REGION Network 29: a | b | c | d | e |
   RUNG wire#powerrail
      I_Contact( #DONE )
      { S7_Templates := "SrcType := WChar" } EQ_Contact(in1 := #UNICODE, in2 := WCHAR#'a')
      Move(in := 16#61, out1 => #ASCII_HEX)
      S_Coil( #DONE )
   END_RUNG
   RUNG wire#powerrail
      I_Contact( #DONE )
      { S7_Templates := "SrcType := WChar" } EQ_Contact(in1 := #UNICODE, in2 := WCHAR#'b')
      Move(in := 16#62, out1 => #ASCII_HEX)
      S_Coil( #DONE )
   END_RUNG
   RUNG wire#powerrail
      I_Contact( #DONE )
      { S7_Templates := "SrcType := WChar" } EQ_Contact(in1 := #UNICODE, in2 := WCHAR#'c')
      Move(in := 16#63, out1 => #ASCII_HEX)
      S_Coil( #DONE )
   END_RUNG
   RUNG wire#powerrail
      I_Contact( #DONE )
      { S7_Templates := "SrcType := WChar" } EQ_Contact(in1 := #UNICODE, in2 := WCHAR#'d')
      Move(in := 16#64, out1 => #ASCII_HEX)
      S_Coil( #DONE )
   END_RUNG
   RUNG wire#powerrail
      I_Contact( #DONE )
      { S7_Templates := "SrcType := WChar" } EQ_Contact(in1 := #UNICODE, in2 := WCHAR#'e')
      Move(in := 16#65, out1 => #ASCII_HEX)
      S_Coil( #DONE )
   END_RUNG
   // the same network as SCL:
   IF NOT #DONE AND (#UNICODE = WCHAR#'a') THEN
       #ASCII_HEX := 16#61;
       #DONE := TRUE;
   END_IF;
   IF NOT #DONE AND (#UNICODE = WCHAR#'b') THEN
       #ASCII_HEX := 16#62;
       #DONE := TRUE;
   END_IF;
   IF NOT #DONE AND (#UNICODE = WCHAR#'c') THEN
       #ASCII_HEX := 16#63;
       #DONE := TRUE;
   END_IF;
   IF NOT #DONE AND (#UNICODE = WCHAR#'d') THEN
       #ASCII_HEX := 16#64;
       #DONE := TRUE;
   END_IF;
   IF NOT #DONE AND (#UNICODE = WCHAR#'e') THEN
       #ASCII_HEX := 16#65;
       #DONE := TRUE;
   END_IF;
END_REGION

REGION Network 30: f | g | h | i | j |
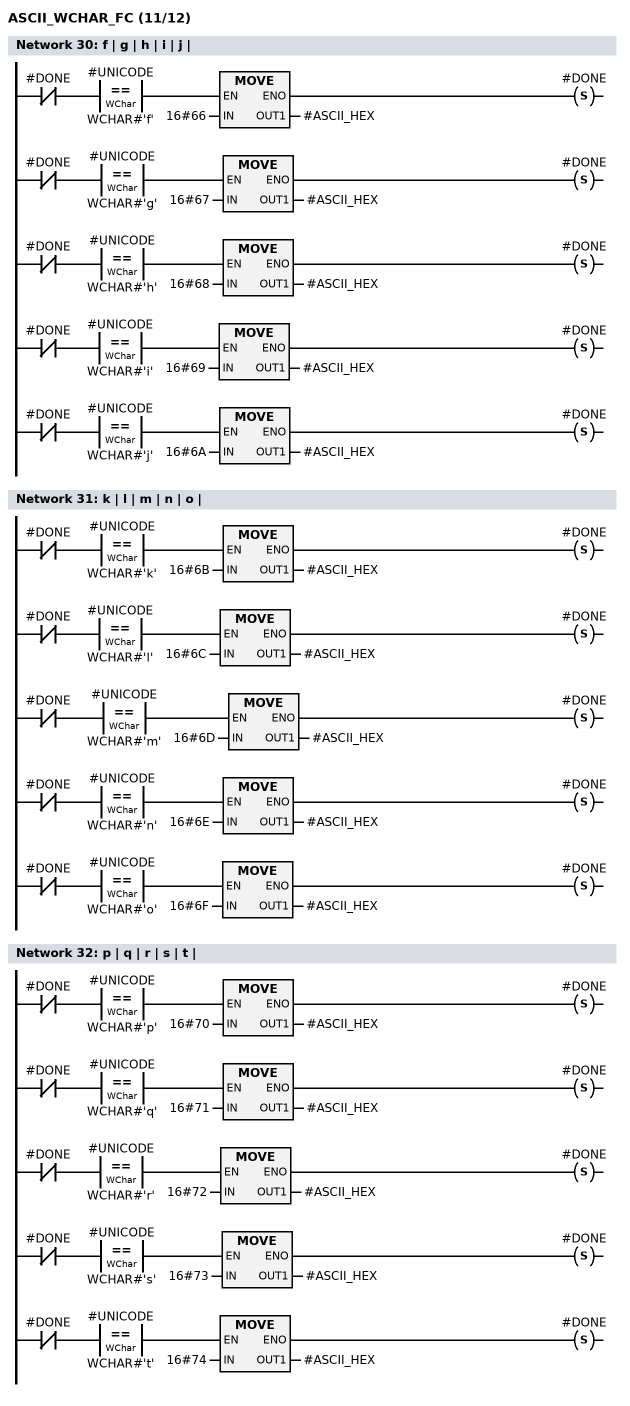
   RUNG wire#powerrail
      I_Contact( #DONE )
      { S7_Templates := "SrcType := WChar" } EQ_Contact(in1 := #UNICODE, in2 := WCHAR#'f')
      Move(in := 16#66, out1 => #ASCII_HEX)
      S_Coil( #DONE )
   END_RUNG
   RUNG wire#powerrail
      I_Contact( #DONE )
      { S7_Templates := "SrcType := WChar" } EQ_Contact(in1 := #UNICODE, in2 := WCHAR#'g')
      Move(in := 16#67, out1 => #ASCII_HEX)
      S_Coil( #DONE )
   END_RUNG
   RUNG wire#powerrail
      I_Contact( #DONE )
      { S7_Templates := "SrcType := WChar" } EQ_Contact(in1 := #UNICODE, in2 := WCHAR#'h')
      Move(in := 16#68, out1 => #ASCII_HEX)
      S_Coil( #DONE )
   END_RUNG
   RUNG wire#powerrail
      I_Contact( #DONE )
      { S7_Templates := "SrcType := WChar" } EQ_Contact(in1 := #UNICODE, in2 := WCHAR#'i')
      Move(in := 16#69, out1 => #ASCII_HEX)
      S_Coil( #DONE )
   END_RUNG
   RUNG wire#powerrail
      I_Contact( #DONE )
      { S7_Templates := "SrcType := WChar" } EQ_Contact(in1 := #UNICODE, in2 := WCHAR#'j')
      Move(in := 16#6A, out1 => #ASCII_HEX)
      S_Coil( #DONE )
   END_RUNG
   // the same network as SCL:
   IF NOT #DONE AND (#UNICODE = WCHAR#'f') THEN
       #ASCII_HEX := 16#66;
       #DONE := TRUE;
   END_IF;
   IF NOT #DONE AND (#UNICODE = WCHAR#'g') THEN
       #ASCII_HEX := 16#67;
       #DONE := TRUE;
   END_IF;
   IF NOT #DONE AND (#UNICODE = WCHAR#'h') THEN
       #ASCII_HEX := 16#68;
       #DONE := TRUE;
   END_IF;
   IF NOT #DONE AND (#UNICODE = WCHAR#'i') THEN
       #ASCII_HEX := 16#69;
       #DONE := TRUE;
   END_IF;
   IF NOT #DONE AND (#UNICODE = WCHAR#'j') THEN
       #ASCII_HEX := 16#6A;
       #DONE := TRUE;
   END_IF;
END_REGION

REGION Network 31: k | l | m | n | o |
   RUNG wire#powerrail
      I_Contact( #DONE )
      { S7_Templates := "SrcType := WChar" } EQ_Contact(in1 := #UNICODE, in2 := WCHAR#'k')
      Move(in := 16#6B, out1 => #ASCII_HEX)
      S_Coil( #DONE )
   END_RUNG
   RUNG wire#powerrail
      I_Contact( #DONE )
      { S7_Templates := "SrcType := WChar" } EQ_Contact(in1 := #UNICODE, in2 := WCHAR#'l')
      Move(in := 16#6C, out1 => #ASCII_HEX)
      S_Coil( #DONE )
   END_RUNG
   RUNG wire#powerrail
      I_Contact( #DONE )
      { S7_Templates := "SrcType := WChar" } EQ_Contact(in1 := #UNICODE, in2 := WCHAR#'m')
      Move(in := 16#6D, out1 => #ASCII_HEX)
      S_Coil( #DONE )
   END_RUNG
   RUNG wire#powerrail
      I_Contact( #DONE )
      { S7_Templates := "SrcType := WChar" } EQ_Contact(in1 := #UNICODE, in2 := WCHAR#'n')
      Move(in := 16#6E, out1 => #ASCII_HEX)
      S_Coil( #DONE )
   END_RUNG
   RUNG wire#powerrail
      I_Contact( #DONE )
      { S7_Templates := "SrcType := WChar" } EQ_Contact(in1 := #UNICODE, in2 := WCHAR#'o')
      Move(in := 16#6F, out1 => #ASCII_HEX)
      S_Coil( #DONE )
   END_RUNG
   // the same network as SCL:
   IF NOT #DONE AND (#UNICODE = WCHAR#'k') THEN
       #ASCII_HEX := 16#6B;
       #DONE := TRUE;
   END_IF;
   IF NOT #DONE AND (#UNICODE = WCHAR#'l') THEN
       #ASCII_HEX := 16#6C;
       #DONE := TRUE;
   END_IF;
   IF NOT #DONE AND (#UNICODE = WCHAR#'m') THEN
       #ASCII_HEX := 16#6D;
       #DONE := TRUE;
   END_IF;
   IF NOT #DONE AND (#UNICODE = WCHAR#'n') THEN
       #ASCII_HEX := 16#6E;
       #DONE := TRUE;
   END_IF;
   IF NOT #DONE AND (#UNICODE = WCHAR#'o') THEN
       #ASCII_HEX := 16#6F;
       #DONE := TRUE;
   END_IF;
END_REGION

REGION Network 32: p | q | r | s | t |
   RUNG wire#powerrail
      I_Contact( #DONE )
      { S7_Templates := "SrcType := WChar" } EQ_Contact(in1 := #UNICODE, in2 := WCHAR#'p')
      Move(in := 16#70, out1 => #ASCII_HEX)
      S_Coil( #DONE )
   END_RUNG
   RUNG wire#powerrail
      I_Contact( #DONE )
      { S7_Templates := "SrcType := WChar" } EQ_Contact(in1 := #UNICODE, in2 := WCHAR#'q')
      Move(in := 16#71, out1 => #ASCII_HEX)
      S_Coil( #DONE )
   END_RUNG
   RUNG wire#powerrail
      I_Contact( #DONE )
      { S7_Templates := "SrcType := WChar" } EQ_Contact(in1 := #UNICODE, in2 := WCHAR#'r')
      Move(in := 16#72, out1 => #ASCII_HEX)
      S_Coil( #DONE )
   END_RUNG
   RUNG wire#powerrail
      I_Contact( #DONE )
      { S7_Templates := "SrcType := WChar" } EQ_Contact(in1 := #UNICODE, in2 := WCHAR#'s')
      Move(in := 16#73, out1 => #ASCII_HEX)
      S_Coil( #DONE )
   END_RUNG
   RUNG wire#powerrail
      I_Contact( #DONE )
      { S7_Templates := "SrcType := WChar" } EQ_Contact(in1 := #UNICODE, in2 := WCHAR#'t')
      Move(in := 16#74, out1 => #ASCII_HEX)
      S_Coil( #DONE )
   END_RUNG
   // the same network as SCL:
   IF NOT #DONE AND (#UNICODE = WCHAR#'p') THEN
       #ASCII_HEX := 16#70;
       #DONE := TRUE;
   END_IF;
   IF NOT #DONE AND (#UNICODE = WCHAR#'q') THEN
       #ASCII_HEX := 16#71;
       #DONE := TRUE;
   END_IF;
   IF NOT #DONE AND (#UNICODE = WCHAR#'r') THEN
       #ASCII_HEX := 16#72;
       #DONE := TRUE;
   END_IF;
   IF NOT #DONE AND (#UNICODE = WCHAR#'s') THEN
       #ASCII_HEX := 16#73;
       #DONE := TRUE;
   END_IF;
   IF NOT #DONE AND (#UNICODE = WCHAR#'t') THEN
       #ASCII_HEX := 16#74;
       #DONE := TRUE;
   END_IF;
END_REGION

REGION Network 33: u | v | w | x | y | z |
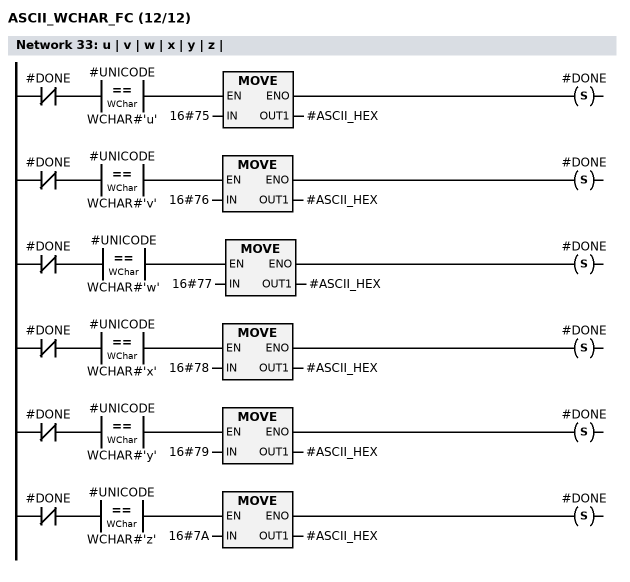
   RUNG wire#powerrail
      I_Contact( #DONE )
      { S7_Templates := "SrcType := WChar" } EQ_Contact(in1 := #UNICODE, in2 := WCHAR#'u')
      Move(in := 16#75, out1 => #ASCII_HEX)
      S_Coil( #DONE )
   END_RUNG
   RUNG wire#powerrail
      I_Contact( #DONE )
      { S7_Templates := "SrcType := WChar" } EQ_Contact(in1 := #UNICODE, in2 := WCHAR#'v')
      Move(in := 16#76, out1 => #ASCII_HEX)
      S_Coil( #DONE )
   END_RUNG
   RUNG wire#powerrail
      I_Contact( #DONE )
      { S7_Templates := "SrcType := WChar" } EQ_Contact(in1 := #UNICODE, in2 := WCHAR#'w')
      Move(in := 16#77, out1 => #ASCII_HEX)
      S_Coil( #DONE )
   END_RUNG
   RUNG wire#powerrail
      I_Contact( #DONE )
      { S7_Templates := "SrcType := WChar" } EQ_Contact(in1 := #UNICODE, in2 := WCHAR#'x')
      Move(in := 16#78, out1 => #ASCII_HEX)
      S_Coil( #DONE )
   END_RUNG
   RUNG wire#powerrail
      I_Contact( #DONE )
      { S7_Templates := "SrcType := WChar" } EQ_Contact(in1 := #UNICODE, in2 := WCHAR#'y')
      Move(in := 16#79, out1 => #ASCII_HEX)
      S_Coil( #DONE )
   END_RUNG
   RUNG wire#powerrail
      I_Contact( #DONE )
      { S7_Templates := "SrcType := WChar" } EQ_Contact(in1 := #UNICODE, in2 := WCHAR#'z')
      Move(in := 16#7A, out1 => #ASCII_HEX)
      S_Coil( #DONE )
   END_RUNG
   // the same network as SCL:
   IF NOT #DONE AND (#UNICODE = WCHAR#'u') THEN
       #ASCII_HEX := 16#75;
       #DONE := TRUE;
   END_IF;
   IF NOT #DONE AND (#UNICODE = WCHAR#'v') THEN
       #ASCII_HEX := 16#76;
       #DONE := TRUE;
   END_IF;
   IF NOT #DONE AND (#UNICODE = WCHAR#'w') THEN
       #ASCII_HEX := 16#77;
       #DONE := TRUE;
   END_IF;
   IF NOT #DONE AND (#UNICODE = WCHAR#'x') THEN
       #ASCII_HEX := 16#78;
       #DONE := TRUE;
   END_IF;
   IF NOT #DONE AND (#UNICODE = WCHAR#'y') THEN
       #ASCII_HEX := 16#79;
       #DONE := TRUE;
   END_IF;
   IF NOT #DONE AND (#UNICODE = WCHAR#'z') THEN
       #ASCII_HEX := 16#7A;
       #DONE := TRUE;
   END_IF;
END_REGION
END_FUNCTION

FUNCTION "INT_TO_WSTRING" : Void   // FC202, SCL
{ S7_Optimized_Access := 'TRUE' }
VERSION : 0.1
   VAR_INPUT
      Value : Int;
      BASE : Array[0..9] of WChar;
      AsTime : Bool;
   END_VAR
   VAR_OUTPUT
      "String" : WString;
   END_VAR
   VAR_TEMP
      x1 : Int;
      x10 : Int;
      x100 : Int;
      x1000 : Int;
      x10000 : Int;
      void : WString[1];
   END_VAR
BEGIN
   #x10000 := #Value / 10000;
   #x1000 := (#Value - #x10000*10000) / 1000;
   #x100 := (#Value - #x10000*10000 - #x1000*1000) / 100;
   #x10 := (#Value - #x10000*10000- #x1000*1000 - #x100*100) / 10;
   #x1 := (#Value - #x10000 * 10000 - #x1000 * 1000 - #x100 * 100 - #x10 * 10) / 1;

   #String := #void;
   IF #x10000 > 0 THEN
       #String := CONCAT_WSTRING(IN1 := #String, IN2 := #BASE[#x10000]);
   END_IF;

   IF #x1000 > 0 THEN
       #String := CONCAT_WSTRING(IN1 := #String, IN2 := #BASE[#x1000]);
   ELSE
       IF #x10000 > 0 THEN
           #String := CONCAT_WSTRING(IN1 := #String, IN2 := #BASE[#x1000]);
       END_IF;
   END_IF;

   IF #x100 > 0 THEN
       #String := CONCAT_WSTRING(IN1 := #String, IN2 := #BASE[#x100]);
   ELSE
       IF #x1000 > 0 OR #x10000 > 0 THEN
           #String := CONCAT_WSTRING(IN1 := #String, IN2 := #BASE[#x100]);
       END_IF;
   END_IF;

   IF #x10 > 0 THEN
       #String := CONCAT_WSTRING(IN1 := #String, IN2 := #BASE[#x10]);
   ELSE
       IF #x100 > 0 OR #x1000 > 0 OR #x10000 > 0 OR #AsTime THEN
           #String := CONCAT_WSTRING(IN1 := #String, IN2 := #BASE[#x10]);
       END_IF;
   END_IF;

   IF #x1 > 0 THEN
       #String := CONCAT_WSTRING(IN1 := #String, IN2 := #BASE[#x1]);
   ELSE
       IF #x10 > 0 OR #x100 > 0 OR #x1000 > 0 OR #x10000 > 0 OR #AsTime THEN
           #String := CONCAT_WSTRING(IN1 := #String, IN2 := #BASE[#x1]);
       END_IF;
   END_IF;
END_FUNCTION

(* ===== HMI "HMI_RT_1" =====
system functions are stored by id; their names below are inferred from use
connection "HMI_Connection_1": ETHERNET, SMART_S7_1200_OMS

HMI tags "Sys"
   "DI_set" : Int AT %DB1.DBW0
   "AI_set" : Int AT %DB1.DBW0
   "DO_set" : Int AT %DB1.DBW0
   "Dos_set" : Int AT %DB1.DBW0
   "AO_Set" : Int AT %DB1.DBW0
   "SP_set" : Int AT %DB1.DBW0
   "Line_set" : Int AT %DB1.DBW0
   "Lines_Alarms" : Int AT %DB1.DBW0
   "MainScr" : Int AT %DB1.DBW0
   "settings" : Int, internal
   "Reset_All" : Bool = PLC Reset_All AT %M3.0, 1 s
   "Alm_Any" : Bool = PLC Alm_Any AT %M15.7, 1 s
   "Time_SYS_DB_RD_Time" : DTL = PLC Time_SYS_DB.RD_Time AT %DB95.DBX130.0, 1 s
   "Time_SYS_DB_SP_Time" : DTL = PLC Time_SYS_DB.SP_Time AT %DB95.DBX142.0, 1 s
   "Hand" : Bool AT %DB1.DBX0.0
   "Sett_scr" : Int AT %DB1.DBX0.0
   "Time_SYS_DB_Set_Time" : Bool = PLC Time_SYS_DB.Set_Time AT %DB95.DBX0.0, 1 s
   "Events" : Word = PLC Events AT %MW200, 1 s
   "Time_SYS_DB_Time_Now_Day" : Int = PLC Time_SYS_DB.Time_Now.Day AT %DB95.DBW6, 1 s
   "Time_SYS_DB_Time_Now_Month" : Int = PLC Time_SYS_DB.Time_Now.Month AT %DB95.DBW4, 1 s
   "Time_SYS_DB_Time_Now_Weekday" : Int = PLC Time_SYS_DB.Time_Now.Weekday AT %DB95.DBW8, 1 s
   "Lines" : Int AT %DB1.DBW0
   "Support_DB_All_AIs" : Int = PLC Support_DB.All_AIs, 1 s
   "Support_DB_All_AOs" : Int = PLC Support_DB.All_AOs, 1 s
   "Support_DB_All_DIs" : Int = PLC Support_DB.All_DIs, 1 s
   "Support_DB_All_DOs" : Int = PLC Support_DB.All_DOs, 1 s
   "Support_DB_DTR_Clean" : Bool = PLC Support_DB.DTR_Clean, 1 s
   "FB_DRV_Start_DB_s1_hour" : Int = PLC FB_DRV_Start_DB.s1_hour, 1 s
   "FB_DRV_Start_DB_s1_minutes" : Int = PLC FB_DRV_Start_DB.s1_minutes, 1 s
   "FB_DRV_Start_DB_s2_hour" : Int = PLC FB_DRV_Start_DB.s2_hour, 1 s
   "FB_DRV_Start_DB_s2_minutes" : Int = PLC FB_DRV_Start_DB.s2_minutes, 1 s
   "Local_Mode" : Bool = PLC Local_Mode AT %M4.0, 1 s
   "Support_DB_All_MDAs" : Int = PLC Support_DB.All_MDAs, 1 s
   "Support_DB_All_MDs" : Int = PLC Support_DB.All_MDs, 1 s
   "Support_DB_All_PIDs" : Int = PLC Support_DB.All_PIDs, 1 s
   "Support_DB_All_VD2s" : Int = PLC Support_DB.All_VD2s, 1 s

HMI tags "Indirect"
   "Vx" : Int AT %DB1.DBW0
   "Vx_Name" : WString[15] AT %DB1.DBW0
   "V_x_Alarms" : Word AT %DB0.DBW50, 1 s
   "V_x_CMD_Force" : Bool AT %DB0.DBX4.7, 1 s
   "V_x_CMD_Hand" : Bool AT %DB0.DBX4.2, 1 s
   "V_x_CMD_Local" : Bool AT %DB0.DBX4.3, 1 s
   "V_x_CMD_Lock" : Bool AT %DB0.DBX4.4, 1 s
   "V_x_CMD_Open" : Bool AT %DB0.DBX2.6, 1 s
   "V_x_CMD_Service" : Bool AT %DB0.DBX4.5, 1 s
   "V_x_CMD_Sim" : Bool AT %DB0.DBX5.2, 1 s
   "V_x_CMD_Start_A" : Bool AT %DB0.DBX4.0, 1 s
   "V_x_CMD_Start_M" : Bool AT %DB0.DBX4.1, 1 s
   "V_x_FB_Close" : Bool AT %DB0.DBX12.4, 1 s
   "V_x_FB_KM_Close" : Bool AT %DB0.DBX12.2, 1 s
   "V_x_FB_KM_Open" : Bool AT %DB0.DBX12.1, 1 s
   "V_x_FB_Open" : Bool AT %DB0.DBX12.3, 1 s
   "V_x_Indirect_BIT_CMD_Close" : Int AT %DB0.DBW96, 1 s
   "V_x_Indirect_BIT_CMD_Open" : Int AT %DB0.DBW94, 1 s
   "V_x_Indirect_BIT_FB_Close" : Int AT %DB0.DBW92, 1 s
   "V_x_Indirect_BIT_FB_Open" : Int AT %DB0.DBW90, 1 s
   "V_x_Indirect_BIT_FB_QF" : Int AT %DB0.DBW84, 1 s
   "V_x_Indirect_BYTE_CMD_Close" : Int AT %DB0.DBW80, 1 s
   "V_x_Indirect_BYTE_CMD_Open" : Int AT %DB0.DBW78, 1 s
   "V_x_Indirect_BYTE_FB_Close" : Int AT %DB0.DBW76, 1 s
   "V_x_Indirect_BYTE_FB_Open" : Int AT %DB0.DBW74, 1 s
   "V_x_Indirect_BYTE_FB_QF" : Int AT %DB0.DBW68, 1 s
   "V_x_Inv_Close" : Bool AT %DB0.DBX46.6, 1 s
   "V_x_Inv_Open" : Bool AT %DB0.DBX46.5, 1 s
   "V_x_Status" : Int AT %DB0.DBW8, 1 s
   "V_x_Use_Close" : Bool AT %DB0.DBX10.4, 1 s
   "V_x_Wait_Off_Now" : Int AT %DB0.DBW30, 1 s
   "V_x_Wait_Off_SP" : Int AT %DB0.DBW28, 1 s
   "V_x_Wait_On_Now" : Int AT %DB0.DBW36, 1 s
   "V_x_Wait_On_SP" : Int AT %DB0.DBW34, 1 s
   "V_x_Use_Open" : Bool AT %DB0.DBX10.3, 1 s
   "M_x_Alarms" : Word AT %DB0.DBW44, 1 s
   "M_x_CMD_Force" : Bool AT %DB0.DBX4.7, 1 s
   "M_x_CMD_Hand" : Bool AT %DB0.DBX4.2, 1 s
   "M_x_CMD_Lock" : Bool AT %DB0.DBX4.4, 1 s
   "M_x_CMD" : Bool AT %DB0.DBX2.3, 1 s
   "M_x_CMD_Start_A" : Bool AT %DB0.DBX4.0, 1 s
   "M_x_CMD_Start_M" : Bool AT %DB0.DBX4.1, 1 s
   "M_x_FB_KM" : Bool AT %DB0.DBX12.1, 1 s
   "M_x_FB_QF" : Bool AT %DB0.DBX12.0, 1 s
   "M_x_Indirect_BIT_CMD" : Int AT %DB0.DBW84, 1 s
   "M_x_Indirect_BIT_FB_KM" : Int AT %DB0.DBW82, 1 s
   "M_x_Indirect_BIT_FB_QF" : Int AT %DB0.DBW80, 1 s
   "M_x_Indirect_BYTE_CMD" : Int AT %DB0.DBW78, 1 s
   "M_x_Indirect_BYTE_FB_KM" : Int AT %DB0.DBW76, 1 s
   "M_x_Indirect_BYTE_FB_QF" : Int AT %DB0.DBW74, 1 s
   "M_x_Indirect_CMD" : Bool AT %DB0.DBX72.2, 1 s
   "M_x_Indirect_FB_KM" : Bool AT %DB0.DBX72.1, 1 s
   "M_x_Indirect_FB_QF" : Bool AT %DB0.DBX72.0, 1 s
   "M_x_Inv_KM" : Bool AT %DB0.DBX40.2, 1 s
   "M_x_Inv_QF" : Bool AT %DB0.DBX40.1, 1 s
   "M_x_OpTime_All_h" : DInt AT %DB0.DBD50, 1 s
   "M_x_Status" : Int AT %DB0.DBW8, 1 s
   "M_x_Use_KM" : Bool AT %DB0.DBX10.1, 1 s
   "M_x_Use_QF" : Bool AT %DB0.DBX10.0, 1 s
   "M_x_Wait_Off_Now" : Int AT %DB0.DBW36, 1 s
   "M_x_Wait_Off_SP" : Int AT %DB0.DBW34, 1 s
   "M_x_Wait_On_Now" : Int AT %DB0.DBW30, 1 s
   "M_x_Wait_On_SP" : Int AT %DB0.DBW28, 1 s
   "MA_x_Converter_Max_In" : Real AT %DB0.DBD114, 1 s
   "MA_x_Converter_Max_Out" : Real AT %DB0.DBD118, 1 s
   "MA_x_Converter_Min_In" : Real AT %DB0.DBD106, 1 s
   "MA_x_Converter_Min_Out" : Real AT %DB0.DBD110, 1 s
   "MA_x_Indirect_BYTE_SP" : Int AT %DB0.DBW94, 1 s
   "Mx" : Int AT %DB1.DBW0
   "Mx_Name" : WString[16] AT %DB1.DBX0.0
   "AIx_Name" : WString[15], internal
   "AIx" : Int, internal
   "AI_x_ADDR" : Int AT %DB0.DBW200, 1 s
   "AI_x_Alarms" : Word AT %DB0.DBW188, 1 s
   "AI_x_Alarm_H" : Bool AT %DB0.DBX186.2, 1 s
   "AI_x_Alarm_HH" : Bool AT %DB0.DBX186.1, 1 s
   "AI_x_Alarm_L" : Bool AT %DB0.DBX186.3, 1 s
   "AI_x_Alarm_LL" : Bool AT %DB0.DBX186.4, 1 s
   "AI_x_Alarm_NC" : Bool AT %DB0.DBX186.5, 1 s
   "AI_x_Alarm_SC" : Bool AT %DB0.DBX186.6, 1 s
   "AI_x_Calibration" : Real AT %DB0.DBD24, 1 s
   "AI_x_CMD_Alarm" : Bool AT %DB0.DBX9.0, 1 s
   "AI_x_CMD_Hand" : Bool AT %DB0.DBX8.2, 1 s
   "AI_x_Converter_Max_In" : Real AT %DB0.DBD46, 1 s
   "AI_x_Converter_Max_Out" : Real AT %DB0.DBD50, 1 s
   "AI_x_Converter_Min_In" : Real AT %DB0.DBD38, 1 s
   "AI_x_Converter_Min_Out" : Real AT %DB0.DBD42, 1 s
   "AI_x_Result" : Real AT %DB0.DBD4, 1 s
   "AI_x_Signal" : Int AT %DB0.DBW2, 1 s
   "AI_x_SP_H" : Real AT %DB0.DBD66, 1 s
   "AI_x_SP_HH" : Real AT %DB0.DBD62, 1 s
   "AI_x_SP_L" : Real AT %DB0.DBD70, 1 s
   "AI_x_SP_LL" : Real AT %DB0.DBD74, 1 s
   "AI_x_Timers_H_SP" : Real AT %DB0.DBD132, 1 s
   "AI_x_Timers_HH_SP" : Real AT %DB0.DBD114, 1 s
   "AI_x_Timers_L_SP" : Real AT %DB0.DBD150, 1 s
   "AI_x_Timers_LL_SP" : Real AT %DB0.DBD168, 1 s
   "AI_x_Use_Filter" : Bool AT %DB0.DBX14.1, 1 s
   "DIx" : Int AT %DB1.DBW0
   "DIx_ADDR_Bit_x_1" : Int AT %DB0.DBW10, 1 s
   "DIx_ADDR_Bit_x_10" : Int AT %DB0.DBW190, 1 s
   "DIx_ADDR_Bit_x_11" : Int AT %DB0.DBW210, 1 s
   "DIx_ADDR_Bit_x_12" : Int AT %DB0.DBW230, 1 s
   "DIx_ADDR_Bit_x_2" : Int AT %DB0.DBW30, 1 s
   "DIx_ADDR_Bit_x_3" : Int AT %DB0.DBW50, 1 s
   "DIx_ADDR_Bit_x_4" : Int AT %DB0.DBW70, 1 s
   "DIx_ADDR_Bit_x_5" : Int AT %DB0.DBW90, 1 s
   "DIx_ADDR_Bit_x_6" : Int AT %DB0.DBW110, 1 s
   "DIx_ADDR_Bit_x_7" : Int AT %DB0.DBW130, 1 s
   "DIx_ADDR_Bit_x_8" : Int AT %DB0.DBW150, 1 s
   "DIx_ADDR_Bit_x_9" : Int AT %DB0.DBW170, 1 s
   "DIx_ADDR_Byte_x_1" : Int AT %DB0.DBW8, 1 s
   "DIx_ADDR_Byte_x_10" : Int AT %DB0.DBW188, 1 s
   "DIx_ADDR_Byte_x_11" : Int AT %DB0.DBW208, 1 s
   "DIx_ADDR_Byte_x_12" : Int AT %DB0.DBW228, 1 s
   "DIx_ADDR_Byte_x_2" : Int AT %DB0.DBW28, 1 s
   "DIx_ADDR_Byte_x_3" : Int AT %DB0.DBW48, 1 s
   "DIx_ADDR_Byte_x_4" : Int AT %DB0.DBW68, 1 s
   "DIx_ADDR_Byte_x_5" : Int AT %DB0.DBW88, 1 s
   "DIx_ADDR_Byte_x_6" : Int AT %DB0.DBW108, 1 s
   "DIx_ADDR_Byte_x_7" : Int AT %DB0.DBW128, 1 s
   "DIx_ADDR_Byte_x_8" : Int AT %DB0.DBW148, 1 s
   "DIx_ADDR_Byte_x_9" : Int AT %DB0.DBW168, 1 s
   "DIx_Hand_x_1" : Bool AT %DB0.DBX4.2, 1 s
   "DIx_Hand_x_10" : Bool AT %DB0.DBX184.2, 1 s
   "DIx_Hand_x_11" : Bool AT %DB0.DBX204.2, 1 s
   "DIx_Hand_x_12" : Bool AT %DB0.DBX224.2, 1 s
   "DIx_Hand_x_2" : Bool AT %DB0.DBX24.2, 1 s
   "DIx_Hand_x_3" : Bool AT %DB0.DBX44.2, 1 s
   "DIx_Hand_x_4" : Bool AT %DB0.DBX64.2, 1 s
   "DIx_Hand_x_5" : Bool AT %DB0.DBX84.2, 1 s
   "DIx_Hand_x_6" : Bool AT %DB0.DBX104.2, 1 s
   "DIx_Hand_x_7" : Bool AT %DB0.DBX124.2, 1 s
   "DIx_Hand_x_8" : Bool AT %DB0.DBX144.2, 1 s
   "DIx_Hand_x_9" : Bool AT %DB0.DBX164.2, 1 s
   "DIx_Inverse_x_1" : Bool AT %DB0.DBX6.0, 1 s
   "DIx_Inverse_x_10" : Bool AT %DB0.DBX186.0, 1 s
   "DIx_Inverse_x_11" : Bool AT %DB0.DBX206.0, 1 s
   "DIx_Inverse_x_12" : Bool AT %DB0.DBX226.0, 1 s
   "DIx_Inverse_x_2" : Bool AT %DB0.DBX26.0, 1 s
   "DIx_Inverse_x_3" : Bool AT %DB0.DBX46.0, 1 s
   "DIx_Inverse_x_4" : Bool AT %DB0.DBX66.0, 1 s
   "DIx_Inverse_x_5" : Bool AT %DB0.DBX86.0, 1 s
   "DIx_Inverse_x_6" : Bool AT %DB0.DBX106.0, 1 s
   "DIx_Inverse_x_7" : Bool AT %DB0.DBX126.0, 1 s
   "DIx_Inverse_x_8" : Bool AT %DB0.DBX146.0, 1 s
   "DIx_Inverse_x_9" : Bool AT %DB0.DBX166.0, 1 s
   "DIx_Start_M_x_1" : Bool AT %DB0.DBX4.1, 1 s
   "DIx_Start_M_x_10" : Bool AT %DB0.DBX184.1, 1 s
   "DIx_Start_M_x_11" : Bool AT %DB0.DBX204.1, 1 s
   "DIx_Start_M_x_12" : Bool AT %DB0.DBX224.1, 1 s
   "DIx_Start_M_x_2" : Bool AT %DB0.DBX24.1, 1 s
   "DIx_Start_M_x_3" : Bool AT %DB0.DBX44.1, 1 s
   "DIx_Start_M_x_4" : Bool AT %DB0.DBX64.1, 1 s
   "DIx_Start_M_x_5" : Bool AT %DB0.DBX84.1, 1 s
   "DIx_Start_M_x_6" : Bool AT %DB0.DBX104.1, 1 s
   "DIx_Start_M_x_7" : Bool AT %DB0.DBX124.1, 1 s
   "DIx_Start_M_x_8" : Bool AT %DB0.DBX144.1, 1 s
   "DIx_Start_M_x_9" : Bool AT %DB0.DBX164.1, 1 s
   "DOx" : Int, internal
   "DOx_ADDR_Bit_x_1" : Int AT %DB0.DBW10, 1 s
   "DOx_ADDR_Bit_x_10" : Int AT %DB0.DBW190, 1 s
   "DOx_ADDR_Bit_x_11" : Int AT %DB0.DBW210, 1 s
   "DOx_ADDR_Bit_x_12" : Int AT %DB0.DBW230, 1 s
   "DOx_ADDR_Bit_x_2" : Int AT %DB0.DBW30, 1 s
   "DOx_ADDR_Bit_x_3" : Int AT %DB0.DBW50, 1 s
   "DOx_ADDR_Bit_x_4" : Int AT %DB0.DBW70, 1 s
   "DOx_ADDR_Bit_x_5" : Int AT %DB0.DBW90, 1 s
   "DOx_ADDR_Bit_x_6" : Int AT %DB0.DBW110, 1 s
   "DOx_ADDR_Bit_x_7" : Int AT %DB0.DBW130, 1 s
   "DOx_ADDR_Bit_x_8" : Int AT %DB0.DBW150, 1 s
   "DOx_ADDR_Bit_x_9" : Int AT %DB0.DBW170, 1 s
   "DOx_ADDR_Byte_x_1" : Int AT %DB0.DBW8, 1 s
   "DOx_ADDR_Byte_x_10" : Int AT %DB0.DBW188, 1 s
   "DOx_ADDR_Byte_x_11" : Int AT %DB0.DBW208, 1 s
   "DOx_ADDR_Byte_x_12" : Int AT %DB0.DBW228, 1 s
   "DOx_ADDR_Byte_x_2" : Int AT %DB0.DBW28, 1 s
   "DOx_ADDR_Byte_x_3" : Int AT %DB0.DBW48, 1 s
   "DOx_ADDR_Byte_x_4" : Int AT %DB0.DBW68, 1 s
   "DOx_ADDR_Byte_x_5" : Int AT %DB0.DBW88, 1 s
   "DOx_ADDR_Byte_x_6" : Int AT %DB0.DBW108, 1 s
   "DOx_ADDR_Byte_x_7" : Int AT %DB0.DBW128, 1 s
   "DOx_ADDR_Byte_x_8" : Int AT %DB0.DBW148, 1 s
   "DOx_ADDR_Byte_x_9" : Int AT %DB0.DBW168, 1 s
   "DOx_Hand_x_1" : Bool AT %DB0.DBX4.2, 1 s
   "DOx_Hand_x_10" : Bool AT %DB0.DBX184.2, 1 s
   "DOx_Hand_x_11" : Bool AT %DB0.DBX204.2, 1 s
   "DOx_Hand_x_12" : Bool AT %DB0.DBX224.2, 1 s
   "DOx_Hand_x_2" : Bool AT %DB0.DBX24.2, 1 s
   "DOx_Hand_x_3" : Bool AT %DB0.DBX44.2, 1 s
   "DOx_Hand_x_4" : Bool AT %DB0.DBX64.2, 1 s
   "DOx_Hand_x_5" : Bool AT %DB0.DBX84.2, 1 s
   "DOx_Hand_x_6" : Bool AT %DB0.DBX104.2, 1 s
   "DOx_Hand_x_7" : Bool AT %DB0.DBX124.2, 1 s
   "DOx_Hand_x_8" : Bool AT %DB0.DBX144.2, 1 s
   "DOx_Hand_x_9" : Bool AT %DB0.DBX164.2, 1 s
   "DOx_Inverse_x_1" : Bool AT %DB0.DBX6.0, 1 s
   "DOx_Inverse_x_10" : Bool AT %DB0.DBX186.0, 1 s
   "DOx_Inverse_x_11" : Bool AT %DB0.DBX206.0, 1 s
   "DOx_Inverse_x_12" : Bool AT %DB0.DBX226.0, 1 s
   "DOx_Inverse_x_2" : Bool AT %DB0.DBX26.0, 1 s
   "DOx_Inverse_x_3" : Bool AT %DB0.DBX46.0, 1 s
   "DOx_Inverse_x_4" : Bool AT %DB0.DBX66.0, 1 s
   "DOx_Inverse_x_5" : Bool AT %DB0.DBX86.0, 1 s
   "DOx_Inverse_x_6" : Bool AT %DB0.DBX106.0, 1 s
   "DOx_Inverse_x_7" : Bool AT %DB0.DBX126.0, 1 s
   "DOx_Inverse_x_8" : Bool AT %DB0.DBX146.0, 1 s
   "DOx_Inverse_x_9" : Bool AT %DB0.DBX166.0, 1 s
   "DOx_Start_M_x_1" : Bool AT %DB0.DBX4.1, 1 s
   "DOx_Start_M_x_10" : Bool AT %DB0.DBX184.1, 1 s
   "DOx_Start_M_x_11" : Bool AT %DB0.DBX204.1, 1 s
   "DOx_Start_M_x_12" : Bool AT %DB0.DBX224.1, 1 s
   "DOx_Start_M_x_2" : Bool AT %DB0.DBX24.1, 1 s
   "DOx_Start_M_x_3" : Bool AT %DB0.DBX44.1, 1 s
   "DOx_Start_M_x_4" : Bool AT %DB0.DBX64.1, 1 s
   "DOx_Start_M_x_5" : Bool AT %DB0.DBX84.1, 1 s
   "DOx_Start_M_x_6" : Bool AT %DB0.DBX104.1, 1 s
   "DOx_Start_M_x_7" : Bool AT %DB0.DBX124.1, 1 s
   "DOx_Start_M_x_8" : Bool AT %DB0.DBX144.1, 1 s
   "DOx_Start_M_x_9" : Bool AT %DB0.DBX164.1, 1 s
   "V_x_CMD_Close" : Bool AT %DB0.DBX2.7, 1 s
   "V_x_Use_Electro" : Bool AT %DB0.DBX10.6, 1 s
   "V_x_Use_Cross" : Bool AT %DB0.DBX10.7, 1 s
   "V_x_Use_CMD_Close" : Bool AT %DB0.DBX11.1, 1 s
   "V_x_Use_CMD_Open" : Bool AT %DB0.DBX11.0, 1 s
   "V_x_Use_QF" : Bool AT %DB0.DBX10.0, 1 s
   "V_x_FB_QF" : Bool AT %DB0.DBX12.0, 1 s
   "V_x_Inv_QF" : Bool AT %DB0.DBX46.1, 1 s
   "M_x_CMD_ResetOpTime" : Bool AT %DB0.DBX5.4, 1 s
   "M_x_OpTime_Now_h" : DInt AT %DB0.DBD62, 1 s
   "M_x_OpTime_SP_h" : DInt AT %DB0.DBD58, 1 s
   "M_x_Use_OpTime" : Bool AT %DB0.DBX10.2, 1 s
   "M_x_OpTime_Alarm" : Bool AT %DB0.DBX42.7, 1 s
   "AI_x_Filter_SP" : Int AT %DB0.DBW202, 1 s
   "M_x_CMD_Local" : Bool AT %DB0.DBX4.3, 1 s
   "AI_x_CMD_Reset" : Bool AT %DB0.DBX9.1, 1 s
   "M_x_CMD_Reset" : Bool AT %DB0.DBX5.1, 1 s
   "V_x_CMD_Reset" : Bool AT %DB0.DBX5.1, 1 s
   "AI_x_Status" : Int AT %DB0.DBW12, 1 s
   "AI_x_VmA" : Real AT %DB0.DBD16, 1 s
   "AI_x_CMD_Start_A" : Bool AT %DB0.DBX8.0, 1 s
   "AI_x_Alarm_ST" : Bool AT %DB0.DBX186.0, 1 s
   "AI_x_Type" : Int AT %DB0.DBW198, 1 s
   "AI_x_Input_Type" : Int AT %DB0.DBW194, 1 s
   "AI_x_CMD_Reset_1" : Bool AT %DB0.DBX9.1, 1 s
   "AI_x_Use_Status" : Bool AT %DB0.DBX14.4, 1 s
   "AI_x_Use_RTD" : Bool AT %DB0.DBX14.0, 1 s
   "AOx_Name" : WString[10], internal
   "AOx" : Int, internal
   "AO_x_ADDR" : Int AT %DB0.DBW60, 1 s
   "AO_x_CMD_Hand" : Bool AT %DB0.DBX8.2, 1 s
   "AO_x_CMD_Start_A" : Bool AT %DB0.DBX8.0, 1 s
   "AO_x_Converter_Max_In" : Real AT %DB0.DBD42, 1 s
   "AO_x_Converter_Max_Out" : Real AT %DB0.DBD46, 1 s
   "AO_x_Converter_Min_In" : Real AT %DB0.DBD34, 1 s
   "AO_x_Converter_Min_Out" : Real AT %DB0.DBD38, 1 s
   "AO_x_Output_Type" : Int AT %DB0.DBW54, 1 s
   "AO_x_Signal" : Int AT %DB0.DBW6, 1 s
   "AO_x_Slow_Step_Down" : Real AT %DB0.DBD76, 1 s
   "AO_x_Slow_Step_Up" : Real AT %DB0.DBD72, 1 s
   "AO_x_Slow_T_Down_SP" : Real AT %DB0.DBD98, 1 s
   "AO_x_Slow_T_Up_SP" : Real AT %DB0.DBD80, 1 s
   "AO_x_Slow_Use_Down" : Bool AT %DB0.DBX70.1, 1 s
   "AO_x_Slow_Use_Up" : Bool AT %DB0.DBX70.0, 1 s
   "AO_x_SP_M" : Real AT %DB0.DBD20, 1 s
   "AO_x_Status" : Int AT %DB0.DBW12, 1 s
   "AO_x_Type" : Int AT %DB0.DBW58, 1 s
   "AO_x_VmA" : Real AT %DB0.DBD16, 1 s
   "M_x_Inv_CMD" : Bool AT %DB0.DBX40.0, 1 s
   "M_x_Delay_On_SP" : Int AT %DB0.DBW22, 1 s
   "M_x_Delay_On_Now" : Int AT %DB0.DBW24, 1 s
   "M_x_Delay_Off_SP" : Int AT %DB0.DBW16, 1 s
   "M_x_Delay_Off_Now" : Int AT %DB0.DBW18, 1 s
   "M_x_CMD_Sim" : Bool AT %DB0.DBX5.2, 1 s
   "V_x_Inv_CMD" : Bool AT %DB0.DBX46.0, 1 s
   "V_x_Delay_Off_Now" : Int AT %DB0.DBW18, 1 s
   "V_x_Delay_Off_SP" : Int AT %DB0.DBW16, 1 s
   "V_x_Delay_On_Now" : Int AT %DB0.DBW24, 1 s
   "V_x_Delay_On_SP" : Int AT %DB0.DBW22, 1 s
   "AI_x_RTD_c" : Real AT %DB0.DBD20, 1 s
   "MA_x_Type" : Int AT %DB0.DBW128, 1 s
   "MA_x_Output_Type" : Int AT %DB0.DBW126, 1 s
   "MA_x_VmA" : Real AT %DB0.DBD122, 1 s
   "MA_x_SP_M" : Real AT %DB0.DBD90, 1 s
   "M_x_CMD_Service" : Bool AT %DB0.DBX4.5, 1 s
   "PIDx" : Int, internal
   "PIDx_Name" : WString[15], internal
   "PID_x_CMD_Start_A" : Bool AT %DB0.DBX16.0, 1 s
   "PID_x_CMD_Hand" : Bool AT %DB0.DBX16.2, 1 s
   "PID_x_CMD_Reset" : Bool AT %DB0.DBX17.1, 1 s
   "PID_x_CMD_Alarm" : Bool AT %DB0.DBX17.0, 1 s
   "PID_x_CMD_Vector" : Bool AT %DB0.DBX17.3, 1 s
   "PID_x_SP_M" : Real AT %DB0.DBD18, 1 s
   "PID_x_PID_Hand" : Real AT %DB0.DBD46, 1 s
   "PID_x_Settings_SP_P" : Real AT %DB0.DBD66, 1 s
   "PID_x_Settings_SP_Ti" : Real AT %DB0.DBD70, 1 s
   "PID_x_Settings_SP_Td" : Real AT %DB0.DBD74, 1 s
   "PID_x_Settings_DeadBand" : Real AT %DB0.DBD106, 1 s
   "PID_x_C_SP" : Real AT %DB0.DBD78, 1 s
   "PID_x_Settings_Max_SP" : Real AT %DB0.DBD82, 1 s
   "PID_x_Settings_Min_SP" : Real AT %DB0.DBD86, 1 s
   "PID_x_Settings_Max_in" : Real AT %DB0.DBD90, 1 s
   "PID_x_Settings_Min_in" : Real AT %DB0.DBD94, 1 s
   "PID_x_Settings_Max_out" : Real AT %DB0.DBD98, 1 s
   "PID_x_Settings_Min_out" : Real AT %DB0.DBD102, 1 s
   "PID_x_Settings_SP_Cycle" : Real AT %DB0.DBD78, 1 s
   "PID_x_x" : Real AT %DB0.DBD26, 1 s
   "PID_x_Value" : Real AT %DB0.DBD6, 1 s
   "PID_x_CMD_Force" : Bool AT %DB0.DBX16.7, 1 s
   "PID_x_Sys_Alm_SP_H" : Bool AT %DB0.DBX50.1, 1 s
   "PID_x_Sys_Alm_SP_L" : Bool AT %DB0.DBX50.2, 1 s
   "PID_x_Sys_Alm_In_H" : Bool AT %DB0.DBX50.3, 1 s
   "PID_x_Sys_Alm_In_L" : Bool AT %DB0.DBX50.4, 1 s
   "PID_x_Sys_Error_code" : DWord AT %DB0.DBD52, 1 s

discrete alarms
   411: 'СБРОС АВАРИЙ', class Warnings, trigger "Events" bit 2
   410: 'АВАРИЙНЫЙ СТОП --- ОТЖАТ', class Warnings, trigger "Events" bit 1
   409: 'АВАРИЙНЫЙ СТОП --- НАЖАТ', class Warnings, trigger "Events" bit 0
   3: 'Аварии сброшены', class Warnings, trigger "Events" bit 2
   1: 'Нажата кнопка аварийного останова', class Warnings, trigger "Events" bit 0
   2: 'Отжата кнопка аварийного останова', class Warnings, trigger "Events" bit 1
   4: 'Все устройства переведены в авторежим', class Warnings, trigger "Events" bit 3

text list "WeekDay": 1 'Понедельник'; 2 'Вторник'; 3 'Среда'; 4 'Четверг'; 5 'Пятница'; 6 'Суббота'; 7 'Воскресенье'

text list "NAME": 0 'Установка приготовления'; 1 'Установка приготовления Ф 1'; 2 'Установка приготовления Ф 2'; 3 'Установка приготовления ПАУ 1'; 4 'Установка приготовления ПАУ 2'; 5 'Установка приготовления соды'; 6 'Установка приготовления СА'

text list "OFF_ON": 0 'Выкл.'; 1 'Вкл.'

text list "Month": 1 'Январь'; 2 'Февраль'; 3 'Март'; 4 'Апрель'; 5 'Май'; 6 'Июнь'; 7 'Июль'; 8 'Август'; 9 'Сентябрь'; 10 'Октябрь'; 11 'Ноябрь'; 12 'Декабрь'

text list "Mode": 0 'Местный'; 1 'Дистанционный'

text list "Hand": 0 'Авто'; 1 'Ручной'

text list "VmA": 0 '4..20 mA'; 1 '0..20 mA'; 2 '0..10 V'; 3 '0..5 V'; 4 'RTD'

text list "Input_Type": 0 '%'; 1 '°С'; 2 'бар'; 3 'л/ч'; 4 'м3/ч'; 5 'м'; 6 'мм'; 7 'кПа'; 8 'Па'; 9 'ppm'; 10 'мм'; 11 'м3/с'; 12 '-'; 13 '-'; 14 '-'; 15 '-'

text list "Output_Type": 0 '%'; 1 'Гц'; 2 'л/ч'; 3 'л/м'; 4 'м3/ч'

text list "VmA_1": 0 '4..20 mA'; 1 '0..20 mA'; 2 '0..10 V'; 3 '0..5 V'

text list "VmA_2": 0 '4..20 mA'; 1 '0..20 mA'; 2 '0..10 V'; 3 '0..5 V'

text list "Air_V": 0 'Без фиксации'; 1 'С фиксацией'

graphic list "Alarm": 0 'no_alarm_1'; 1 'alarm'

graphic list "check_blue_inverse": 1 'check_box_off'; 0 'check_box_on'

graphic list "Fan": 0 'fan_1'; 1 'REQ_vent_1'; 2..3 'fan_wait'; 4..999 'fan_error'

graphic list "Filter": 0 'Filter_OFF'; 1 'Filter_WAIT'

graphic list "Link": 0 'Link_Ok'; 1 'Link_Error_1'

graphic list "mixer": 0 'void'; 1 'mix_off'; 2 'mix_on'; 3 'mix_on_2'

graphic list "Motor": 0 'm_off_1'; 1 'm_on_1'; 2..3 'm_wait_1'; 4..1000 'm_alarm_1'

graphic list "Motor_h": 0 'm_off_h'; 1 'm_on_h'; 2..3 'm_wait_h'; 5..1000 'm_alarm_h'; 4 'm_serv_h'

graphic list "OFF_ON": 1 'off_t'; 0 'on_t'

graphic list "check_blue": 0 'check_box_off'; 1 'check_box_on'

graphic list "check_green": 0 'check_box_off'; 1 'ON_Box'

graphic list "Pump_D": 0 'p_off1'; 1 'p_on1'; 2..3 'p_wait1'; 4..1000 'p_alarm1'

graphic list "Pump_L": 0 'p_off'; 1 'p_on'; 2..3 'p_wait'; 4..1000 'p_alarm'

graphic list "Pump_R": 0 'p_off_r'; 1 'p_on_r_3'; 2..3 'p_wait_r'; 4..1000 'p_alarm_r'

graphic list "Pump_U": 0 'P_OFF_Up'; 1 'P_ON_Up'; 2..3 'P_Wait_Up'; 4..1000 'P_Alarm_Up'

graphic list "PIPE_Selector_Green": 0 'void'; 1 'Graphic_8'; 2 'Graphic_10'; 3 'Graphic_5'; 10 'Graphic_31'; 11 'Graphic_37'; 12 'Graphic_36'; 13 'Graphic_12'; 4 'Graphic_33'; 5 'Graphic_6'; 6 'Graphic_41'; 7 'Graphic_35'

graphic list "RT": 0 'RT'; 1 'RT_1'

graphic list "signal_blue": 0 'circle_box_off_1'; 1 'circle_box_on_blue_1'

graphic list "signal_red": 0 'circle_box_off_2'; 1 'circle_box_on_red'

graphic list "Valve_Hor": 0 'v_off'; 1 'v_on'; 2..3 'v_wait'; 4..1000 'v_alarm'

graphic list "Valve_Hor_Analog": 0 'va_off'; 1 'va_on'; 2..3 'va_wait'; 4..1000 'va_alarm'

graphic list "Valve_Vert_L": 0 'v_off4'; 1 'v_on4'; 2..3 'v_wait4'; 4..1000 'v_alarm4'

graphic list "Valve_Vert_R": 0 'v_off2'; 1 'v_on2'; 2..3 'v_wait2'; 4..1000 'v_alarm2'

graphic list "Vent": 0 'mix_off'; 1 'mix_on'; 2..4 'mix_wait_off'; 5..1000 'mix_alarm'

graphic list "Z": 0 'v_c_close'; 1 'v_c_open'; 2..3 'v_c_wait'; 4 'v_c_not'; 5..1000 'v_c_a_1'

graphic list "ON_OFF": 0 'off_t'; 1 'on_t'

graphic list "Local_Mode": 0 'local'; 1 'link_offx'

graphic list "Turn_ON": 0 'off_t'; 1 'on_t'

graphic list "ok_green": 0 'check_box_off'; 1 'ON_Box'

graphic list "signal_green": 0 'circle_box_off_1'; 1 'circle_box_on_green'

graphic list "signal_green_1": 0 'circle_box_off_2'; 1 'circle_box_on_green'

Template "Main" 800x480
   Button "Button_5" at 735,275 size 60x60; TextOff 'Text'; PictureOff "home_1"; PictureList "Alarm"
      on Click: ActivateScreen("Alarms", 0); SetTag("MainScr", 4); SetTag("Support_DB_DTR_Clean", 0)
      Appearance <- "MainScr"
      ProcessValue <- "Alm_Any"
   Button "Button_7" at 735,410 size 60x60; TextOff 'Text'; PictureOff "reset"
      on Click: SetBit("Reset_All")
   Button "Button_8" at 735,5 size 60x60; TextOff 'Text'; PictureOff "home_3"
      on Click: ActivateScreen("Root screen", 0); SetTag("MainScr", 0); SetTag("Support_DB_DTR_Clean", 0)
   Button "Button_9" at 735,5 size 60x60; TextOff 'Text'; PictureOff "home_pressed_1"
      on Click: ActivateScreen("Root screen", 0); SetTag("MainScr", 0)
      Visibility <- "MainScr"
   Button "Button_10" at 735,72 size 60x60; TextOff 'Text'; PictureOff "sett"
      on Click: SetTag("MainScr", 1); ActivateScreen("Select_Settings", 0); SetTag("settings", 0); SetTag("Support_DB_DTR_Clean", 0)
   Button "Button_11" at 735,72 size 60x60; TextOff 'Text'; PictureOff "sett_pressed"
      on Click: SetTag("MainScr", 1); ActivateScreen("Select_Settings", 0); SetTag("settings", 0); SetTag("Support_DB_DTR_Clean", 0)
      Visibility <- "MainScr"
   Button "Button_12" at 735,140 size 60x60; TextOff 'Text'; PictureOff "table"
      on Click: SetTag("MainScr", 2); ActivateScreen("Select_Alarms", 0); SetTag("Support_DB_DTR_Clean", 0)
   Button "Button_13" at 735,207 size 60x60; TextOff 'Text'; PictureOff "history"
      on Click: ActivateScreen("Select_History", 0); SetTag("MainScr", 3); SetTag("Support_DB_DTR_Clean", 0)
   Button "Button_15" at 735,140 size 60x60; TextOff 'Text'; PictureOff "table_pressed"
      on Click: SetTag("MainScr", 2); ActivateScreen("Select_Alarms", 0); SetTag("Support_DB_DTR_Clean", 0)
      Visibility <- "MainScr"
   Button "Button_16" at 735,207 size 60x60; TextOff 'Text'; PictureOff "history_pressed"
      on Click: ActivateScreen("Select_History", 0); SetTag("MainScr", 3); SetTag("Support_DB_DTR_Clean", 0)
      Appearance <- "MainScr"
      Visibility <- "MainScr"
   Button "Template_Button_2" at 735,342 size 60x60; TextOff 'Text'; PictureOff "vdk1"
      on Click: ActivateScreen("About", 0); SetTag("Support_DB_DTR_Clean", 0)

screen "About" 800x480, template "Main"
   TextField "Text field_1" at 274,13 size 212x47; Text 'ООО "VDK"'
   TextField "Text field_4" at 66,74 size 661x96; Text 'Компания VDK производит оборудование для широкого спектра технологических процессов в разных областях промышленности, специализируясь на технологиях подготовки, ввода и перемешивания реагентов.'
   TextField "Text field_2" at 35,231 size 354x73; Text 'Контактная информация: Адрес: Россия, г. Москва, 111116 ул. Лефортовский вал, д. 7Г, стр. 5'
   TextField "Text field_3" at 63,342 size 299x27; Text 'Телефон: +7 (495) 763-29-73'
   TextField "Text field_5" at 132,370 size 160x27; Text 'info@vdktech.ru'
   GraphicView "Graphic view_2" at 492,179 size 189x291; Picture "vdk2_1"

screen "Alarms" 800x480, template "Main"
   AlarmView "Alarm view_1" at 4,3 size 718x439; ColumnTextDate 'Дата / Datum'; ColumnTextAlarmState 'Статус / Status'; ColumnTextTime 'Время / Zeit'; ColumnTextAlarmText 'Аварийное сообщение / Text'; AlarmLog "Alarm_log_1"
   DateTimeField "Date/time field_1" at 253,445 size 116x32
   DateTimeField "Date/time field_2" at 364,445 size 111x32
   TextField "Text field_1" at 580,449 size 144x23; Text 'Сброс аварий ->'
   Button "Button_1" at 9,445 size 150x32; TextOff 'К событиям'
      on Click: ActivateScreen("Events", 0); SetTag("MainScr", 4)

screen "Events" 800x480, template "Main"
   AlarmView "Alarm view_1" at 4,3 size 718x439; ColumnTextDate 'Дата / Datum'; ColumnTextAlarmState 'Статус / Status'; ColumnTextTime 'Время / Zeit'; ColumnTextAlarmText 'Событие / Text'; AlarmLog "Alarm_log_1"
   Button "Button_1" at 9,445 size 150x32; TextOff 'К авариям'
      on Click: ActivateScreen("Alarms", 0); SetTag("MainScr", 4)
   DateTimeField "Date/time field_1" at 253,445 size 116x32
   DateTimeField "Date/time field_2" at 364,445 size 111x32

screen "Select_Alarms" 800x480, template "Main"
   TextField "Text field_29" at 281,6 size 234x33; Text 'Настройка аварий'
   Button "Button_4" at 327,73 size 150x32; TextOff 'Авария'
      on Click: SetTag("MainScr", 2)
   TextField "Text field_2" at 342,44 size 87x28; Text 'Участок'

screen "Select_History" 800x480, template "Main"
   TextField "Text field_29" at 265,6 size 226x33; Text 'Недельный отчёт'
   TextField "Text field_2" at 10,418 size 79x23; Text 'Смена 1:'
   TextField "Text field_3" at 10,450 size 79x23; Text 'Смена 2:'
   IOField "I/O field_6" at 124,419 size 30x24; Authorization "User administration"; FormatPattern 99
      ProcessValue <- "FB_DRV_Start_DB_s1_hour"
   TextField "Text field_13" at 160,419 size 25x23; Text 'ч'
   IOField "I/O field_8" at 180,419 size 30x24; Authorization "User administration"; FormatPattern 99
      ProcessValue <- "FB_DRV_Start_DB_s1_minutes"
   TextField "Text field_14" at 216,419 size 25x23; Text 'м'
   IOField "I/O field_1" at 124,451 size 30x24; Authorization "User administration"; FormatPattern 99
      ProcessValue <- "FB_DRV_Start_DB_s2_hour"
   TextField "Text field_15" at 160,451 size 25x23; Text 'ч'
   IOField "I/O field_2" at 180,451 size 30x24; Authorization "User administration"; FormatPattern 99
      ProcessValue <- "FB_DRV_Start_DB_s2_minutes"
   TextField "Text field_16" at 216,451 size 25x23; Text 'м'

screen "Select_Settings" 800x480, template "Settings"
   TextField "Text field_29" at 249,6 size 293x33; Text 'Настройка параметров'
   Button "Button_4" at 321,73 size 150x32; TextOff 'Основные'; Authorization "Operate"
      on Click: SetTag("MainScr", 1)
   TextField "Text field_1" at 346,44 size 103x28; Text 'PolyMix 1'
   TextField "Text field_3" at 125,411 size 150x27; Text 'Режим работы'
   Button "Button_3" at 124,439 size 150x32; TextOff 'Местный'; Authorization "Operate"; TextList "Mode"
      on Click: ResetBit("Local_Mode")
      Appearance <- "Local_Mode"
      ProcessValue <- "Local_Mode"

